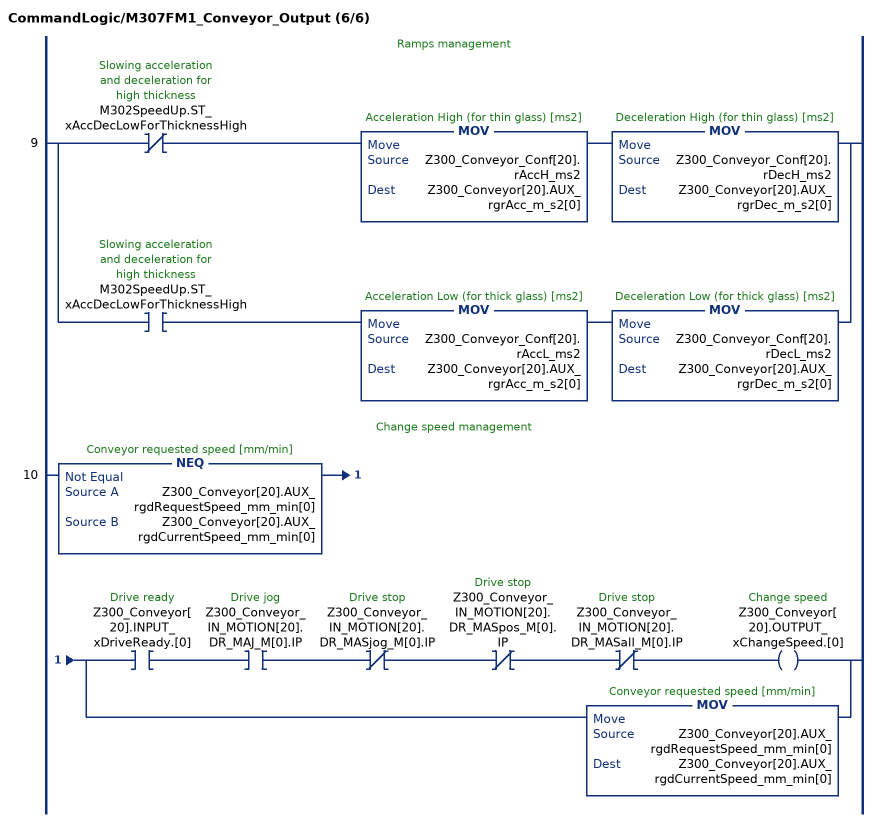
   // Ramps management
   9: [XIO(M302SpeedUp.ST_xAccDecLowForThicknessHigh) MOV(Z300_Conveyor_Conf[20].rAccH_ms2,Z300_Conveyor[20].AUX_rgrAcc_m_s2[0]) MOV(Z300_Conveyor_Conf[20].rDecH_ms2,Z300_Conveyor[20].AUX_rgrDec_m_s2[0]) ,XIC(M302SpeedUp.ST_xAccDecLowForThicknessHigh) MOV(Z300_Conveyor_Conf[20].rAccL_ms2,Z300_Conveyor[20].AUX_rgrAcc_m_s2[0]) MOV(Z300_Conveyor_Conf[20].rDecL_ms2,Z300_Conveyor[20].AUX_rgrDec_m_s2[0]) ];
   // Change speed management
   10: NEQ(Z300_Conveyor[20].AUX_rgdRequestSpeed_mm_min[0],Z300_Conveyor[20].AUX_rgdCurrentSpeed_mm_min[0])[XIC(Z300_Conveyor[20].INPUT_xDriveReady.[0]) XIC(Z300_Conveyor_IN_MOTION[20].DR_MAJ_M[0].IP) XIO(Z300_Conveyor_IN_MOTION[20].DR_MASjog_M[0].IP) XIO(Z300_Conveyor_IN_MOTION[20].DR_MASpos_M[0].IP) XIO(Z300_Conveyor_IN_MOTION[20].DR_MASall_M[0].IP) OTE(Z300_Conveyor[20].OUTPUT_xChangeSpeed.[0]) ,MOV(Z300_Conveyor[20].AUX_rgdRequestSpeed_mm_min[0],Z300_Conveyor[20].AUX_rgdCurrentSpeed_mm_min[0]) ];
END_ROUTINE

ROUTINE M310B_Output   (* ladder *)
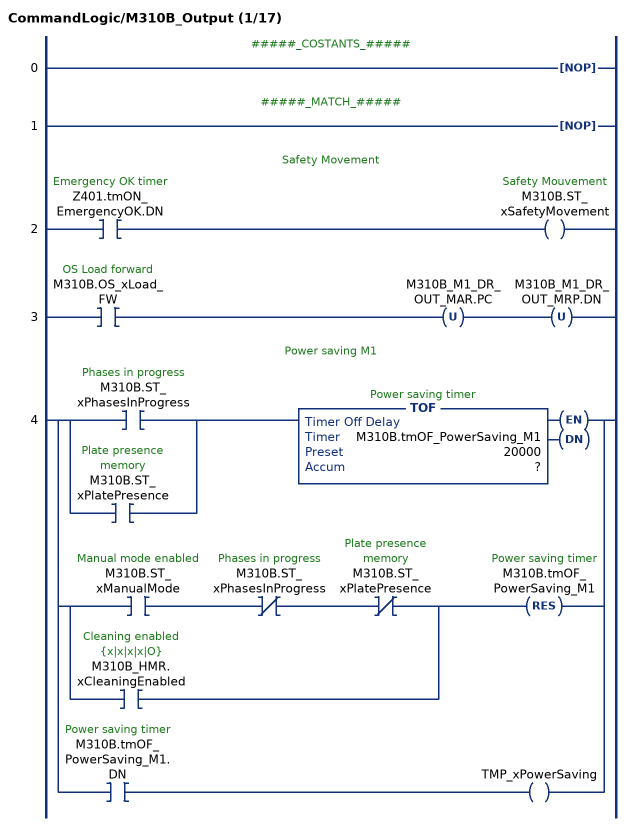
   // #####_COSTANTS_#####
   0: NOP();
   // #####_MATCH_#####
   1: NOP();
   // Safety Movement
   2: XIC(Z401.tmON_EmergencyOK.DN)OTE(M310B.ST_xSafetyMovement);
   3: XIC(M310B.OS_xLoad_FW)OTU(M310B_M1_DR_OUT_MAR.PC)OTU(M310B_M1_DR_OUT_MRP.DN);
   // Power saving M1
   4: [[XIC(M310B.ST_xPhasesInProgress) ,XIC(M310B.ST_xPlatePresence) ] TOF(M310B.tmOF_PowerSaving_M1,?,?) ,[XIC(M310B.ST_xManualMode) XIO(M310B.ST_xPhasesInProgress) XIO(M310B.ST_xPlatePresence) ,XIC(M310B_HMR.xCleaningEnabled) ] RES(M310B.tmOF_PowerSaving_M1) ,XIC(M310B.tmOF_PowerSaving_M1.DN) OTE(TMP_xPowerSaving) ];
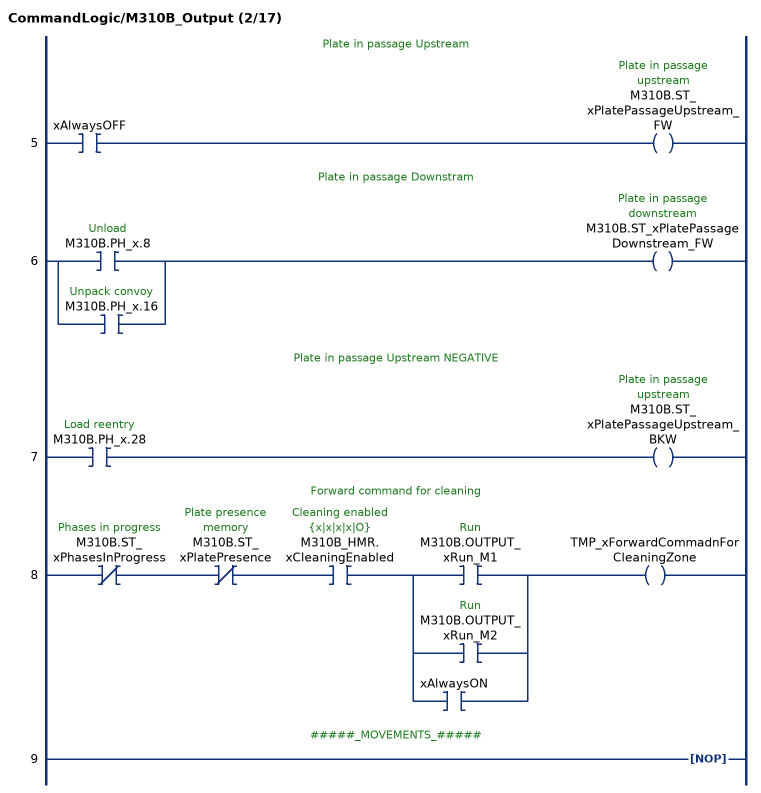
   // Plate in passage Upstream
   5: XIC(xAlwaysOFF)OTE(M310B.ST_xPlatePassageUpstream_FW);
   // Plate in passage Downstram
   6: [XIC(M310B.PH_x.8) ,XIC(M310B.PH_x.16) ]OTE(M310B.ST_xPlatePassageDownstream_FW);
   // Plate in passage Upstream NEGATIVE
   7: XIC(M310B.PH_x.28)OTE(M310B.ST_xPlatePassageUpstream_BKW);
   // Forward command for cleaning
   8: XIO(M310B.ST_xPhasesInProgress)XIO(M310B.ST_xPlatePresence)XIC(M310B_HMR.xCleaningEnabled)[XIC(M310B.OUTPUT_xRun_M1) ,XIC(M310B.OUTPUT_xRun_M2) ,XIC(xAlwaysON) ]OTE(TMP_xForwardCommadnForCleaningZone);
   // #####_MOVEMENTS_#####
   9: NOP();
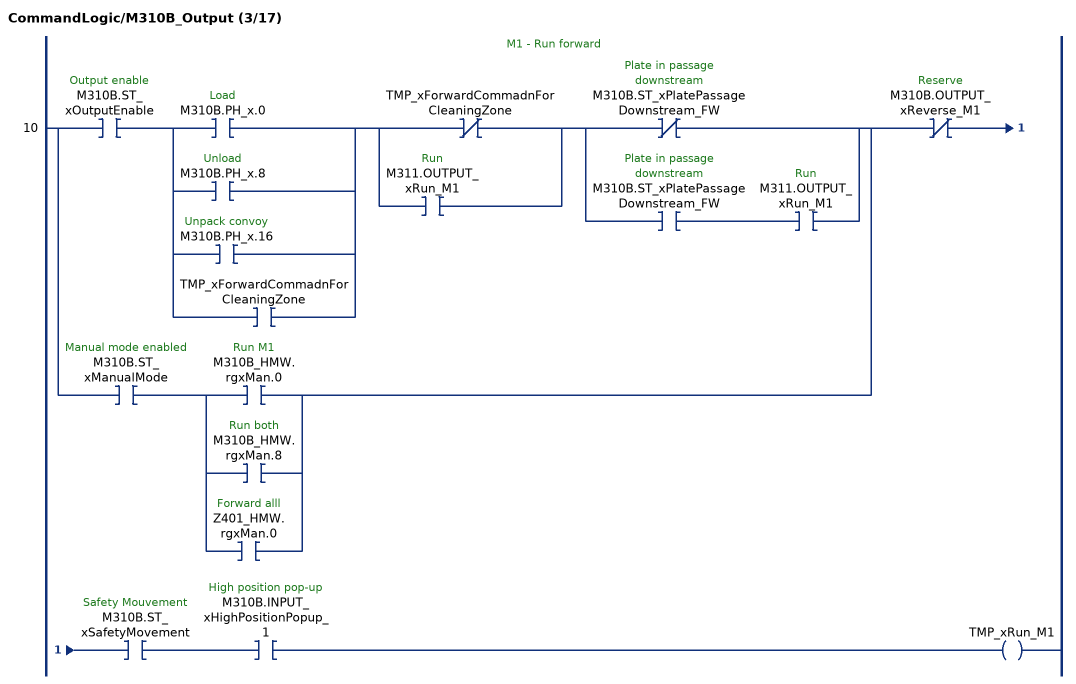
   // M1 - Run forward
   10: [XIC(M310B.ST_xOutputEnable) [XIC(M310B.PH_x.0) ,XIC(M310B.PH_x.8) ,XIC(M310B.PH_x.16) ,XIC(TMP_xForwardCommadnForCleaningZone) ] [XIO(TMP_xForwardCommadnForCleaningZone) ,XIC(M311.OUTPUT_xRun_M1) ] [XIO(M310B.ST_xPlatePassageDownstream_FW) ,XIC(M310B.ST_xPlatePassageDownstream_FW) XIC(M311.OUTPUT_xRun_M1) ] ,XIC(M310B.ST_xManualMode) [XIC(M310B_HMW.rgxMan.0) ,XIC(M310B_HMW.rgxMan.8) ,XIC(Z401_HMW.rgxMan.0) ] ]XIO(M310B.OUTPUT_xReverse_M1)XIC(M310B.ST_xSafetyMovement)XIC(M310B.INPUT_xHighPositionPopup_1)OTE(TMP_xRun_M1);
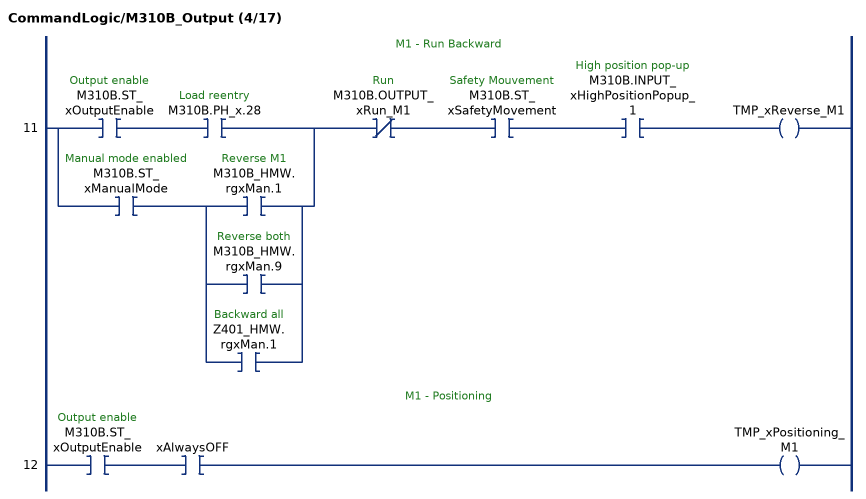
   // M1 - Run Backward
   11: [XIC(M310B.ST_xOutputEnable) XIC(M310B.PH_x.28) ,XIC(M310B.ST_xManualMode) [XIC(M310B_HMW.rgxMan.1) ,XIC(M310B_HMW.rgxMan.9) ,XIC(Z401_HMW.rgxMan.1) ] ]XIO(M310B.OUTPUT_xRun_M1)XIC(M310B.ST_xSafetyMovement)XIC(M310B.INPUT_xHighPositionPopup_1)OTE(TMP_xReverse_M1);
   // M1 - Positioning
   12: XIC(M310B.ST_xOutputEnable)XIC(xAlwaysOFF)OTE(TMP_xPositioning_M1);
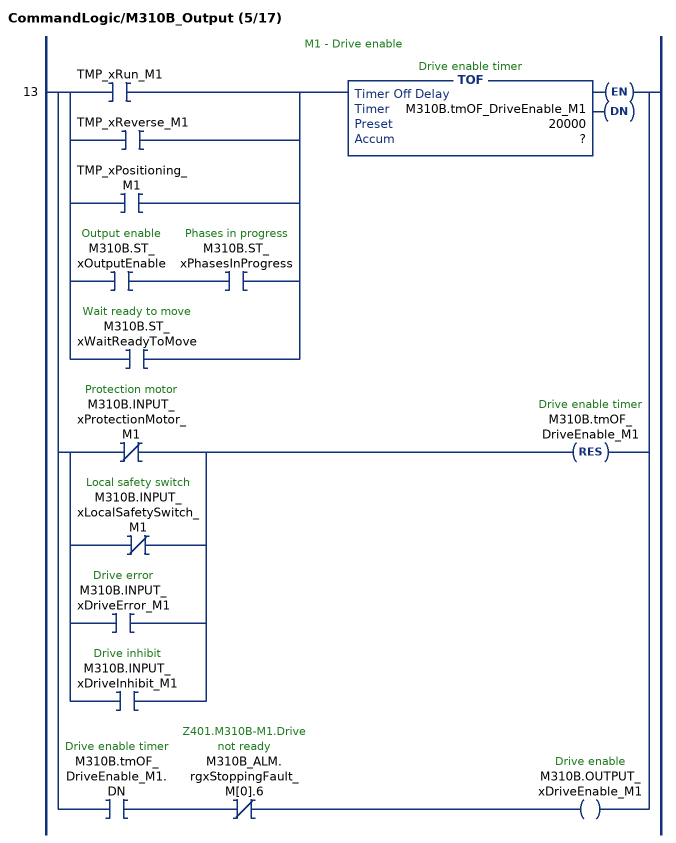
   // M1 - Drive enable
   13: [[XIC(TMP_xRun_M1) ,XIC(TMP_xReverse_M1) ,XIC(TMP_xPositioning_M1) ,XIC(M310B.ST_xOutputEnable) XIC(M310B.ST_xPhasesInProgress) ,XIC(M310B.ST_xWaitReadyToMove) ] TOF(M310B.tmOF_DriveEnable_M1,?,?) ,[XIO(M310B.INPUT_xProtectionMotor_M1) ,XIO(M310B.INPUT_xLocalSafetySwitch_M1) ,XIC(M310B.INPUT_xDriveError_M1) ,XIC(M310B.INPUT_xDriveInhibit_M1) ] RES(M310B.tmOF_DriveEnable_M1) ,XIC(M310B.tmOF_DriveEnable_M1.DN) XIO(M310B_ALM.rgxStoppingFault_M[0].6) OTE(M310B.OUTPUT_xDriveEnable_M1) ];
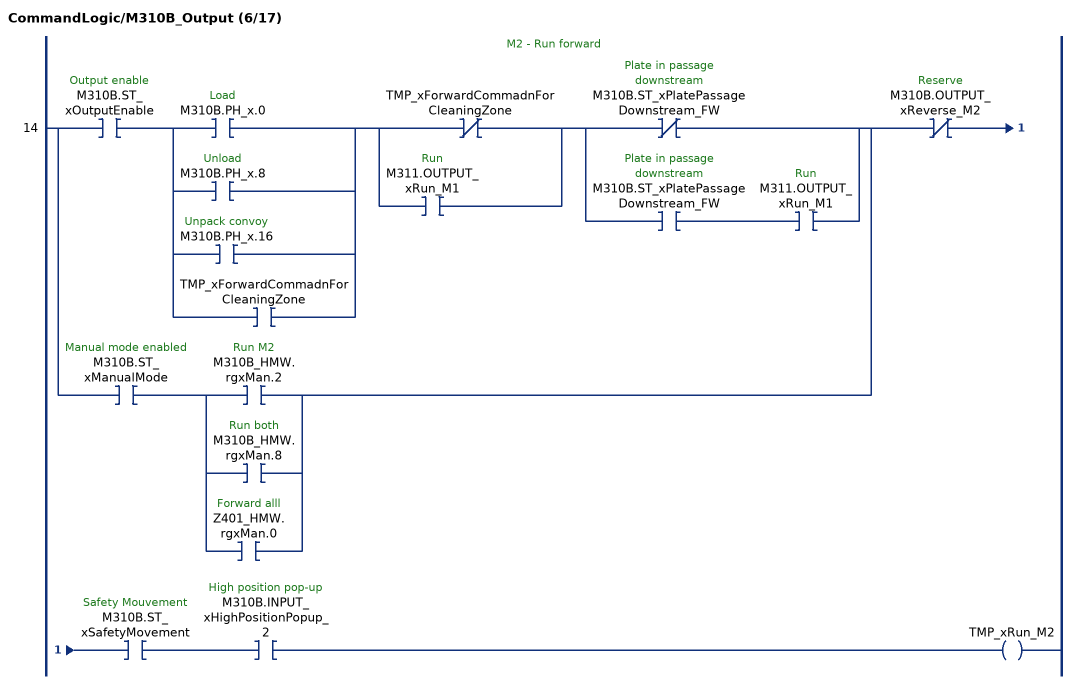
   // M2 - Run forward
   14: [XIC(M310B.ST_xOutputEnable) [XIC(M310B.PH_x.0) ,XIC(M310B.PH_x.8) ,XIC(M310B.PH_x.16) ,XIC(TMP_xForwardCommadnForCleaningZone) ] [XIO(TMP_xForwardCommadnForCleaningZone) ,XIC(M311.OUTPUT_xRun_M1) ] [XIO(M310B.ST_xPlatePassageDownstream_FW) ,XIC(M310B.ST_xPlatePassageDownstream_FW) XIC(M311.OUTPUT_xRun_M1) ] ,XIC(M310B.ST_xManualMode) [XIC(M310B_HMW.rgxMan.2) ,XIC(M310B_HMW.rgxMan.8) ,XIC(Z401_HMW.rgxMan.0) ] ]XIO(M310B.OUTPUT_xReverse_M2)XIC(M310B.ST_xSafetyMovement)XIC(M310B.INPUT_xHighPositionPopup_2)OTE(TMP_xRun_M2);
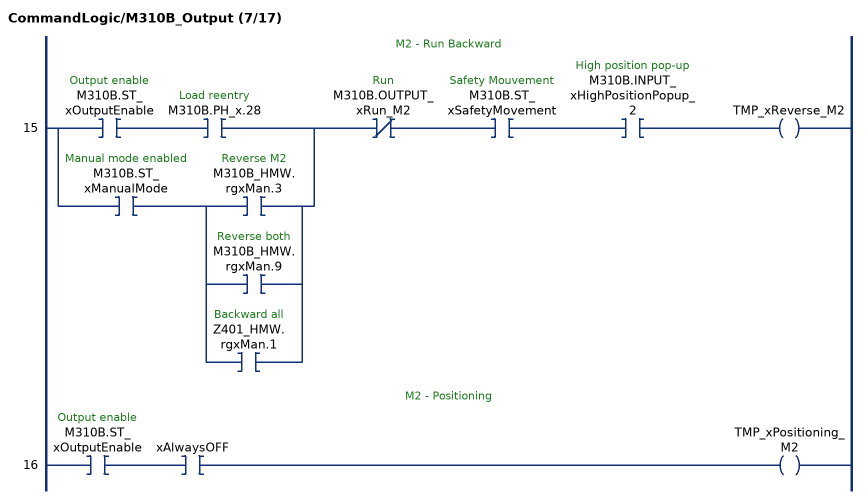
   // M2 - Run Backward
   15: [XIC(M310B.ST_xOutputEnable) XIC(M310B.PH_x.28) ,XIC(M310B.ST_xManualMode) [XIC(M310B_HMW.rgxMan.3) ,XIC(M310B_HMW.rgxMan.9) ,XIC(Z401_HMW.rgxMan.1) ] ]XIO(M310B.OUTPUT_xRun_M2)XIC(M310B.ST_xSafetyMovement)XIC(M310B.INPUT_xHighPositionPopup_2)OTE(TMP_xReverse_M2);
   // M2 - Positioning
   16: XIC(M310B.ST_xOutputEnable)XIC(xAlwaysOFF)OTE(TMP_xPositioning_M2);
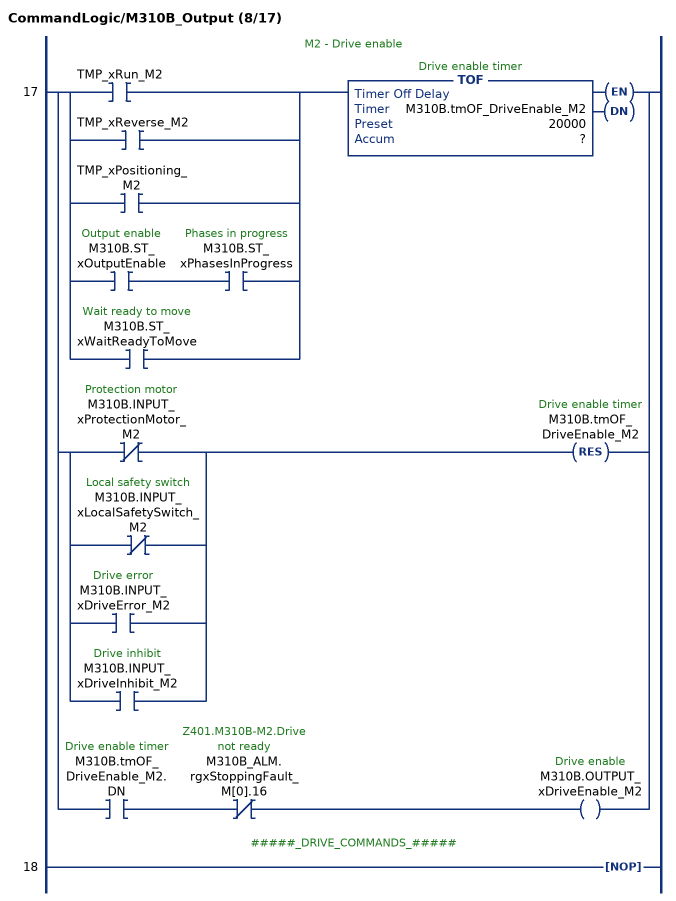
   // M2 - Drive enable
   17: [[XIC(TMP_xRun_M2) ,XIC(TMP_xReverse_M2) ,XIC(TMP_xPositioning_M2) ,XIC(M310B.ST_xOutputEnable) XIC(M310B.ST_xPhasesInProgress) ,XIC(M310B.ST_xWaitReadyToMove) ] TOF(M310B.tmOF_DriveEnable_M2,?,?) ,[XIO(M310B.INPUT_xProtectionMotor_M2) ,XIO(M310B.INPUT_xLocalSafetySwitch_M2) ,XIC(M310B.INPUT_xDriveError_M2) ,XIC(M310B.INPUT_xDriveInhibit_M2) ] RES(M310B.tmOF_DriveEnable_M2) ,XIC(M310B.tmOF_DriveEnable_M2.DN) XIO(M310B_ALM.rgxStoppingFault_M[0].16) OTE(M310B.OUTPUT_xDriveEnable_M2) ];
   // #####_DRIVE_COMMANDS_#####
   18: NOP();
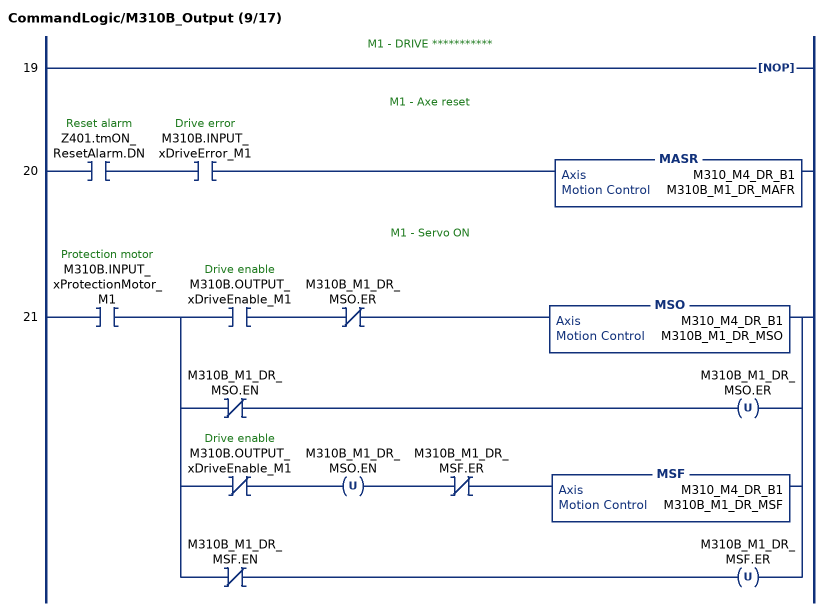
   // M1 - DRIVE ***********
   19: NOP();
   // M1 - Axe reset
   20: XIC(Z401.tmON_ResetAlarm.DN)XIC(M310B.INPUT_xDriveError_M1)MASR(M310_M4_DR_B1,M310B_M1_DR_MAFR);
   // M1 - Servo ON
   21: XIC(M310B.INPUT_xProtectionMotor_M1)[XIC(M310B.OUTPUT_xDriveEnable_M1) XIO(M310B_M1_DR_MSO.ER) MSO(M310_M4_DR_B1,M310B_M1_DR_MSO) ,XIO(M310B_M1_DR_MSO.EN) OTU(M310B_M1_DR_MSO.ER) ,XIO(M310B.OUTPUT_xDriveEnable_M1) OTU(M310B_M1_DR_MSO.EN) XIO(M310B_M1_DR_MSF.ER) MSF(M310_M4_DR_B1,M310B_M1_DR_MSF) ,XIO(M310B_M1_DR_MSF.EN) OTU(M310B_M1_DR_MSF.ER) ];
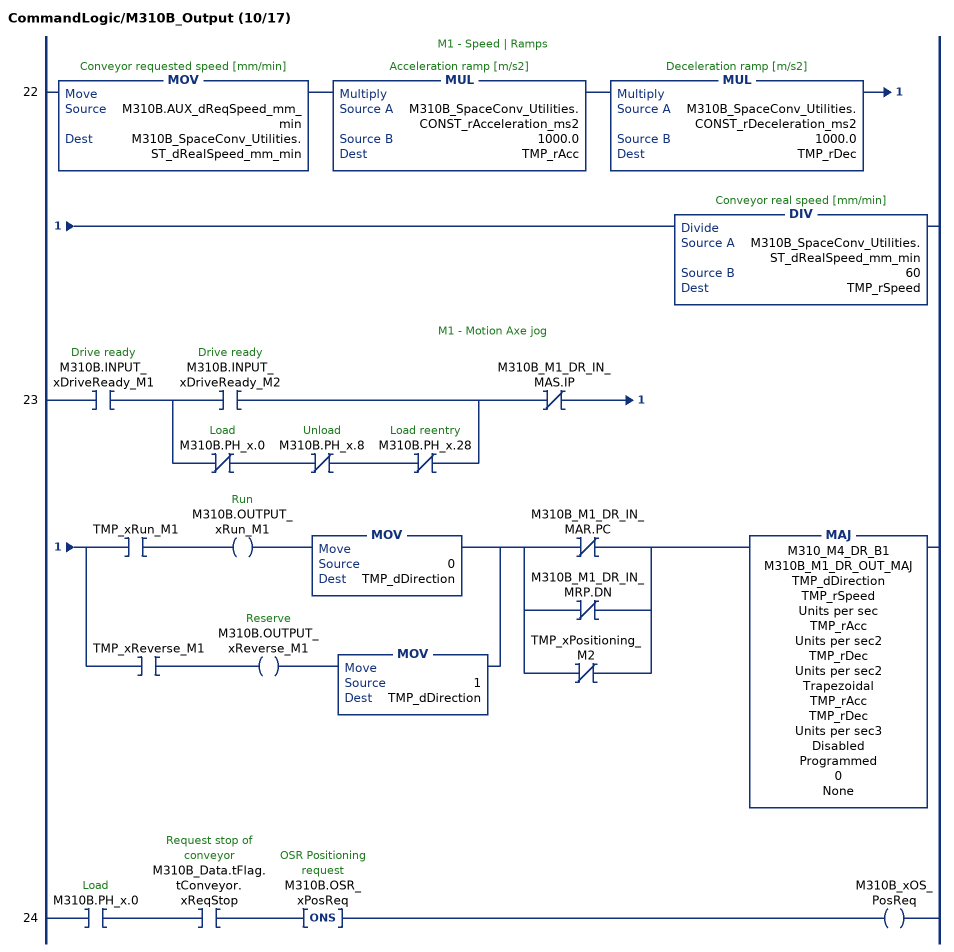
   // M1 - Speed | Ramps
   22: MOV(M310B.AUX_dReqSpeed_mm_min,M310B_SpaceConv_Utilities.ST_dRealSpeed_mm_min)MUL(M310B_SpaceConv_Utilities.CONST_rAcceleration_ms2,1000.0,TMP_rAcc)MUL(M310B_SpaceConv_Utilities.CONST_rDeceleration_ms2,1000.0,TMP_rDec)DIV(M310B_SpaceConv_Utilities.ST_dRealSpeed_mm_min,60,TMP_rSpeed);
   // M1 - Motion Axe jog
   23: XIC(M310B.INPUT_xDriveReady_M1)[XIC(M310B.INPUT_xDriveReady_M2) ,XIO(M310B.PH_x.0) XIO(M310B.PH_x.8) XIO(M310B.PH_x.28) ]XIO(M310B_M1_DR_IN_MAS.IP)[XIC(TMP_xRun_M1) OTE(M310B.OUTPUT_xRun_M1) MOV(0,TMP_dDirection) ,XIC(TMP_xReverse_M1) OTE(M310B.OUTPUT_xReverse_M1) MOV(1,TMP_dDirection) ][XIO(M310B_M1_DR_IN_MAR.PC) ,XIO(M310B_M1_DR_IN_MRP.DN) ,XIO(TMP_xPositioning_M2) ]MAJ(M310_M4_DR_B1,M310B_M1_DR_OUT_MAJ,TMP_dDirection,TMP_rSpeed,Units per sec,TMP_rAcc,Units per sec2,TMP_rDec,Units per sec2,Trapezoidal,TMP_rAcc,TMP_rDec,Units per sec3,Disabled,Programmed,0,None);
   24: XIC(M310B.PH_x.0)XIC(M310B_Data.tFlag.tConveyor.xReqStop)ONS(M310B.OSR_xPosReq)OTE(M310B_xOS_PosReq);
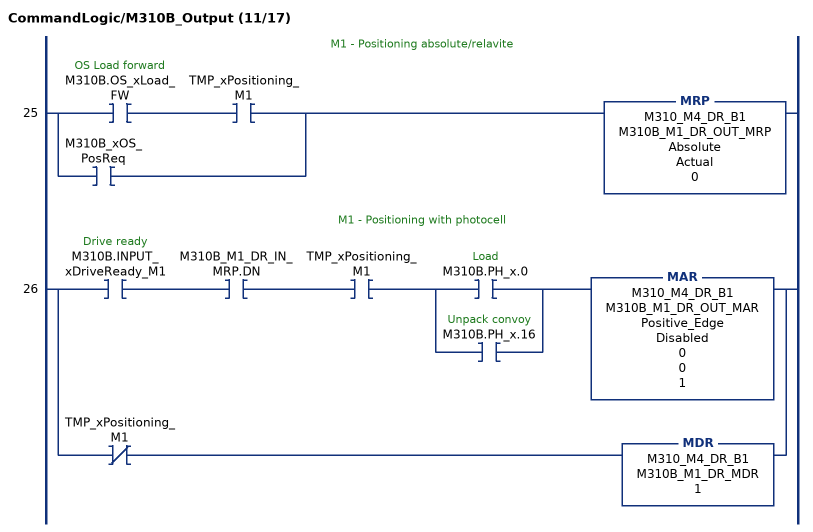
   // M1 - Positioning absolute/relavite
   25: [XIC(M310B.OS_xLoad_FW) XIC(TMP_xPositioning_M1) ,XIC(M310B_xOS_PosReq) ]MRP(M310_M4_DR_B1,M310B_M1_DR_OUT_MRP,Absolute,Actual,0);
   // M1 - Positioning with photocell
   26: [XIC(M310B.INPUT_xDriveReady_M1) XIC(M310B_M1_DR_IN_MRP.DN) XIC(TMP_xPositioning_M1) [XIC(M310B.PH_x.0) ,XIC(M310B.PH_x.16) ] MAR(M310_M4_DR_B1,M310B_M1_DR_OUT_MAR,Positive_Edge,Disabled,0,0,1) ,XIO(TMP_xPositioning_M1) MDR(M310_M4_DR_B1,M310B_M1_DR_MDR,1) ];
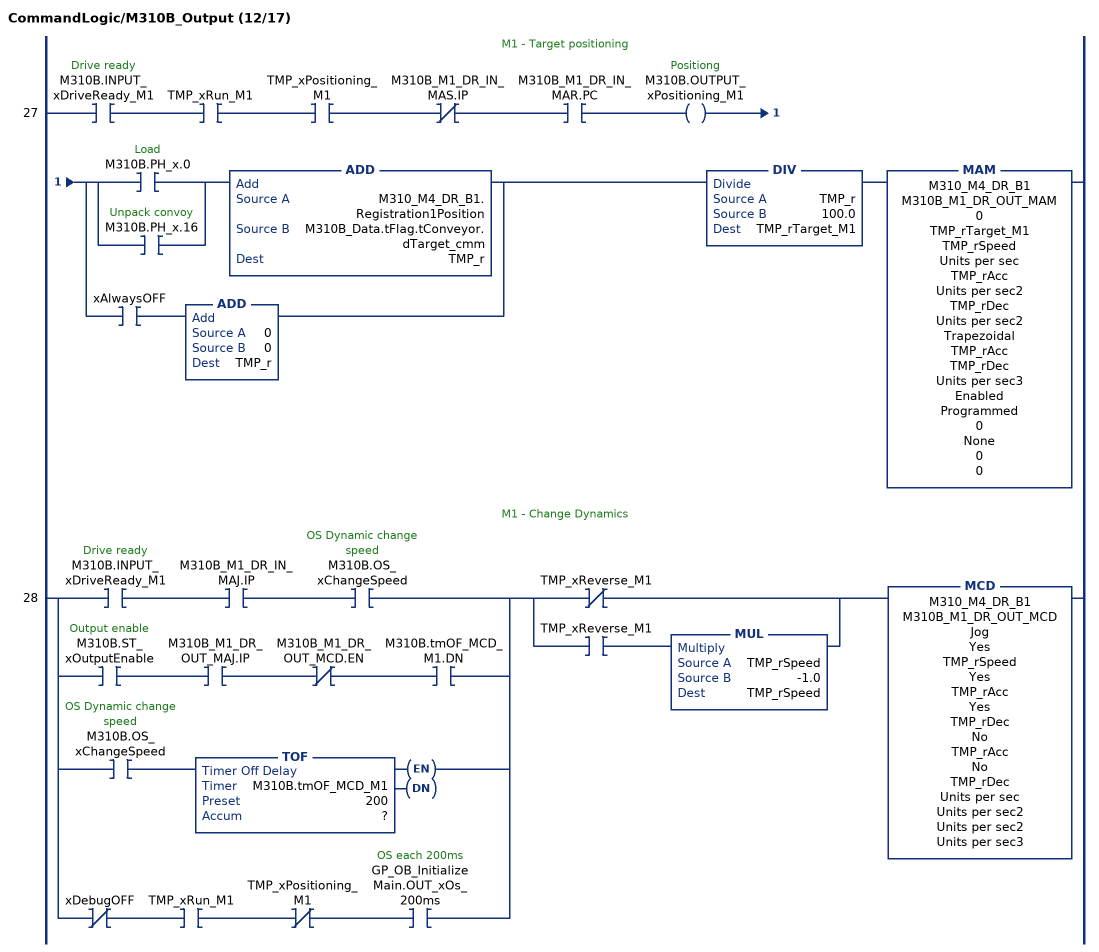
   // M1 - Target positioning
   27: XIC(M310B.INPUT_xDriveReady_M1)XIC(TMP_xRun_M1)XIC(TMP_xPositioning_M1)XIO(M310B_M1_DR_IN_MAS.IP)XIC(M310B_M1_DR_IN_MAR.PC)OTE(M310B.OUTPUT_xPositioning_M1)[[XIC(M310B.PH_x.0) ,XIC(M310B.PH_x.16) ] ADD(M310_M4_DR_B1.Registration1Position,M310B_Data.tFlag.tConveyor.dTarget_cmm,TMP_r) ,XIC(xAlwaysOFF) ADD(0,0,TMP_r) ]DIV(TMP_r,100.0,TMP_rTarget_M1)MAM(M310_M4_DR_B1,M310B_M1_DR_OUT_MAM,0,TMP_rTarget_M1,TMP_rSpeed,Units per sec,TMP_rAcc,Units per sec2,TMP_rDec,Units per sec2,Trapezoidal,TMP_rAcc,TMP_rDec,Units per sec3,Enabled,Programmed,0,None,0,0);
   // M1 - Change Dynamics
   28: [XIC(M310B.INPUT_xDriveReady_M1) XIC(M310B_M1_DR_IN_MAJ.IP) XIC(M310B.OS_xChangeSpeed) ,XIC(M310B.ST_xOutputEnable) XIC(M310B_M1_DR_OUT_MAJ.IP) XIO(M310B_M1_DR_OUT_MCD.EN) XIC(M310B.tmOF_MCD_M1.DN) ,XIC(M310B.OS_xChangeSpeed) TOF(M310B.tmOF_MCD_M1,?,?) ,XIO(xDebugOFF) XIC(TMP_xRun_M1) XIO(TMP_xPositioning_M1) XIC(GP_OB_InitializeMain.OUT_xOs_200ms) ][XIO(TMP_xReverse_M1) ,XIC(TMP_xReverse_M1) MUL(TMP_rSpeed,-1.0,TMP_rSpeed) ]MCD(M310_M4_DR_B1,M310B_M1_DR_OUT_MCD,Jog,Yes,TMP_rSpeed,Yes,TMP_rAcc,Yes,TMP_rDec,No,TMP_rAcc,No,TMP_rDec,Units per sec,Units per sec2,Units per sec2,Units per sec3);
